
ScreenModuleEditorView "ControlMotor-NoAUTO" 640x480
   Button "Botón_1" at 10,10 size 109x37
   Button "Botón_2" at 10,50 size 109x37
   Button "Botón_3" at 130,10 size 101x37
   Button "Botón_4" at 130,50 size 101x37
*)

(* ===== HMI "HMI_RT_1" =====

text list "Enclavamientos": 0 ''; 1 ''; 2 ''; 3 ''; 4 ''; 5 ''

ScreenModuleEditorView "Faceplate_7" 640x480
   Button "Botón_3" at 25,15 size 189x37
   Button "Botón_1" at 11,10 size 93x40
   Button "Botón_2" at 11,54 size 93x40
   IOField "Campo ES_1" at 143,19 size 84x26
   IOField "Campo ES_2" at 143,62 size 84x26
   TextField "Campo de texto_2" at 109,19 size 27x23
   TextField "Campo de texto_3" at 109,62 size 32x23
   IOField "Campo ES_3" at 143,19 size 84x26
   IOField "Campo ES_4" at 143,62 size 84x26
   TextField "Campo de texto_4" at 109,19 size 27x23
   TextField "Campo de texto_5" at 109,62 size 32x23
   TextField "Campo de texto_1" at 10,31 size 97x40
*)

(* ===== HMI "HMI_RT_1" =====

text list "Enclavamientos": 0 ''; 1 ''; 2 ''; 3 ''; 4 ''; 5 ''

ScreenModuleEditorView "Faceplate_2" 640x480
   TextField "Campo de texto_14" at 112,50 size 40x22
   TextField "Campo de texto_13" at 112,14 size 40x22
   TextField "Campo de texto_1" at 67,18 size 125x50
   Button "Botón_1" at 11,10 size 93x32
   Button "Botón_2" at 11,46 size 93x32
   Button "Botón_3" at 136,10 size 117x32
   Button "Botón_4" at 136,46 size 117x32
   SymbolicIOField "Campo ES simbólico_2" at 158,12 size 96x27
   SymbolicIOField "Campo ES simbólico_3" at 158,47 size 96x27
*)

(* ===== HMI "HMI_RT_1" =====

text list "EstadoMotor": 0 ''; 1 ''; 2 ''; 3 ''; 4 ''; 5 ''; 6 ''; 7 ''

ScreenModuleEditorView "ControlMotor-NoAUTO" 640x480
   Button "Botón_1" at 10,10 size 109x37
   Button "Botón_2" at 10,50 size 109x37
   Button "Botón_3" at 130,10 size 101x37
   Button "Botón_4" at 130,50 size 101x37
*)

(* ===== HMI "HMI_RT_1" =====

ScreenModuleEditorView "Faceplate_4" 640x480
   TextField "Campo de texto_14" at 117,50 size 25x22
   TextField "Campo de texto_13" at 119,14 size 23x22
   IOField "Campo ES_9" at 147,48 size 83x29
   IOField "Campo ES_8" at 147,12 size 83x29
   Button "Botón_1" at 10,10 size 93x32
   Button "Botón_2" at 10,46 size 93x32
   Button "Botón_3" at 122,10 size 109x32
   Button "Botón_4" at 122,46 size 109x32
*)

(* ===== HMI "HMI_RT_1" =====

ScreenModuleEditorView "Faceplate_1" 640x480
   TextField "Campo de texto_14" at 117,50 size 25x22
   TextField "Campo de texto_13" at 119,14 size 23x22
   IOField "Campo ES_9" at 147,48 size 83x29
   IOField "Campo ES_8" at 147,12 size 83x29
   Button "Botón_1" at 10,10 size 93x32
   Button "Botón_2" at 10,46 size 93x32
   Button "Botón_3" at 122,10 size 109x32
   Button "Botón_4" at 122,46 size 109x32
*)

(* ===== HMI "HMI_RT_1" =====

ScreenModuleEditorView "Faceplate_1" 640x480
   TextField "Campo de texto_14" at 118,50 size 25x22
   TextField "Campo de texto_13" at 120,14 size 23x22
   TextField "Campo de texto_1" at 59,18 size 125x50
   IOField "Campo ES_9" at 148,48 size 83x29
   IOField "Campo ES_8" at 148,12 size 83x29
   Button "Botón_1" at 11,10 size 93x32
   Button "Botón_2" at 11,46 size 93x32
   Button "Botón_3" at 123,10 size 109x32
   Button "Botón_4" at 123,46 size 109x32
*)

(* ===== HMI "HMI_RT_1" =====

text list "Enclavamientos": 0 ''; 1 ''; 2 ''; 3 ''; 4 ''; 5 ''

ScreenModuleEditorView "Faceplate_10" 640x480
   Button "Botón_3" at 38,10 size 189x37
   Button "Botón_1" at 38,10 size 93x40
   Button "Botón_2" at 133,10 size 93x40
   IOField "Campo ES_1" at 44,75 size 84x26
   IOField "Campo ES_2" at 44,110 size 84x26
   TextField "Campo de texto_2" at 10,75 size 27x23
   TextField "Campo de texto_3" at 10,110 size 32x23
   IOField "Campo ES_3" at 140,75 size 84x26
   IOField "Campo ES_4" at 140,110 size 84x26
   TextField "Campo de texto_4" at 60,51 size 45x23
   TextField "Campo de texto_5" at 146,51 size 71x23
   IOField "Campo ES_5" at 44,75 size 84x26
   IOField "Campo ES_6" at 44,110 size 84x26
   IOField "Campo ES_7" at 140,75 size 84x26
   IOField "Campo ES_8" at 140,110 size 84x26
   TextField "Campo de texto_6" at 10,75 size 27x23
   TextField "Campo de texto_7" at 10,110 size 32x23
   TextField "Campo de texto_8" at 60,51 size 45x23
   TextField "Campo de texto_9" at 146,51 size 71x23
   TextField "Campo de texto_1" at 77,12 size 108x42
*)

(* ===== HMI "HMI_RT_1" =====

ScreenModuleEditorView "Faceplate_6" 640x480
   GraphicIOField "PlotLight_Round_GN" at 52,10 size 35x34
   GraphicIOField "PlotLight_Round_RN" at 10,10 size 34x34
   GraphicView "Visor de gráficos_1" at 52,10 size 34x34
   GraphicView "Visor de gráficos_2" at 53,10 size 34x34
*)

(* ===== HMI "HMI_RT_1" =====

ScreenModuleEditorView "Faceplate_1" 640x480
   Button "Botón_1" at 10,10 size 93x32
   Button "Botón_2" at 10,46 size 93x32
   Button "Botón_3" at 122,10 size 109x32
   Button "Botón_4" at 122,46 size 109x32
*)

(* ===== HMI "HMI_RT_1" =====
connection "Conexión-PLC_2": ETHERNET, SIMATIC S7 300/400 MPI
connection "Conexión-SentronPac_": ETHERNET, MODBUS_TCP

HMI tags "Tabla de variables estándar"
   "IndR6" : Bool, 100 ms
   "IndVparp6" : Bool, 1 s
   "Auto6" : Bool, 1 s
   "PanMCH6" : Bool, 1 s
   "LimSUP6" : Real, 1 s
   "LimINF6" : Real, 1 s
   "VCMP6" : Int, 1 s
   "IncP6" : Bool, 100 ms
   "DecP6" : Bool, 1 s
   "SPONF6" : Real, 1 s
   "SPOFFF6" : Real, 1 s
   "ForzarMarcha6" : Bool, 1 s
   "ForzarParada6" : Bool, 1 s
   "ForzandoMarcha6" : Bool, 1 s
   "SPON6" : Real, 1 s
   "SPOFF6" : Real, 1 s
   "AnimMenuMC006" : Int, 1 s
   "MantMC006" : Bool, 1 s
   "MarchaOK6" : Bool, 1 s
   "MarchaMC006" : Bool, 1 s
   "ParadaMC006" : Bool, 1 s
   "HORAS6" : DInt, 1 s
   "MIN6" : Int, 1 s
   "AnimMotorMC006" : Byte, 1 s
   "EV6" : Bool, 1 s
   "EnclavCompAltaConFlujostato" : Bool = PLC "EnclavCompAltaConFlujostato", 1 s
   "ProxMantMC001_1" : DInt = PLC "ProxMantMC001_1", 1 s
   "ProxMantMC001_2" : DInt = PLC "ProxMantMC001_2", 1 s
   "Varios_UltimoMantMC001_1" : DInt, 1 s
   "Varios_UltimoMantMC001_2" : DInt, 1 s
   "ProxMantMC002_1" : DInt = PLC "ProxMantMC002_1", 1 s
   "ProxMantMC002_2" : DInt = PLC "ProxMantMC002_2", 1 s
   "ProxMantMC003_1" : DInt = PLC "ProxMantMC003_1", 1 s
   "ProxMantMC003_2" : DInt = PLC "ProxMantMC003_2", 1 s
   "ProxMantMC004_1" : DInt = PLC "ProxMantMC004_1", 1 s
   "ProxMantMC004_2" : DInt = PLC "ProxMantMC004_2", 1 s
   "ProxMantMC005_1" : DInt = PLC "ProxMantMC005_1", 1 s
   "ProxMantMC005_2" : DInt = PLC "ProxMantMC005_2", 1 s
   "ProxMantMC006_1" : DInt = PLC "ProxMantMC006_1", 1 s
   "ProxMantMC006_2" : DInt = PLC "ProxMantMC006_2", 1 s
   "Varios_UltimoMantMC002_1" : DInt, 1 s
   "Varios_UltimoMantMC002_2" : DInt, 1 s
   "Varios_UltimoMantMC003_1" : DInt, 1 s
   "Varios_UltimoMantMC003_2" : DInt, 1 s
   "Varios_UltimoMantMC004_1" : DInt, 1 s
   "Varios_UltimoMantMC004_2" : DInt, 1 s
   "Varios_UltimoMantMC005_1" : DInt, 1 s
   "Varios_UltimoMantMC005_2" : DInt, 1 s
   "Varios_UltimoMantMC006_1" : DInt, 1 s
   "Varios_UltimoMantMC006_2" : DInt, 1 s
   "Varios_HorasMantMC001_1" : DInt, 1 s
   "Varios_HorasMantMC006_1" : DInt, 1 s
   "Varios_HorasMantMC006_2" : DInt, 1 s
   "Varios_HorasMantMC002_1" : DInt, 1 s
   "Varios_HorasMantMC001_2" : DInt, 1 s
   "Varios_HorasMantMC002_2" : DInt, 1 s
   "Varios_HorasMantMC004_1" : DInt, 1 s
   "Varios_HorasMantMC004_2" : DInt, 1 s
   "Varios_HorasMantMC005_1" : DInt, 1 s
   "Varios_HorasMantMC005_2" : DInt, 1 s
   "Varios_HorasMantMC003_1" : DInt, 1 s
   "Varios_HorasMantMC003_2" : DInt, 1 s
   "EstadoMantMC003" : Byte = PLC "EstadoMantMC003", 1 s
   "EstadoMantMC005" : Byte = PLC "EstadoMantMC005", 1 s
   "EstadoMantMC004" : Byte = PLC "EstadoMantMC004", 1 s
   "EstadoMantMC002" : Byte = PLC "EstadoMantMC002", 1 s
   "EstadoMantMC001" : Byte = PLC "EstadoMantMC001", 1 s
   "EstadoMantMC006" : Byte = PLC "EstadoMantMC006", 1 s
   "LimiteMantMC001_1" : Bool = PLC "LimiteMantMC001_1", 1 s
   "LimiteMantMC001_2" : Bool = PLC "LimiteMantMC001_2", 1 s
   "LimiteMantMC002_1" : Bool = PLC "LimiteMantMC002_1", 1 s
   "LimiteMantMC002_2" : Bool = PLC "LimiteMantMC002_2", 1 s
   "LimiteMantMC003_1" : Bool = PLC "LimiteMantMC003_1", 1 s
   "LimiteMantMC003_2" : Bool = PLC "LimiteMantMC003_2", 1 s
   "LimiteMantMC004_1" : Bool = PLC "LimiteMantMC004_1", 1 s
   "LimiteMantMC004_2" : Bool = PLC "LimiteMantMC004_2", 1 s
   "LimiteMantMC005_1" : Bool = PLC "LimiteMantMC005_1", 1 s
   "LimiteMantMC005_2" : Bool = PLC "LimiteMantMC005_2", 1 s
   "LimiteMantMC006_1" : Bool = PLC "LimiteMantMC006_1", 1 s
   "LimiteMantMC006_2" : Bool = PLC "LimiteMantMC006_2", 1 s
   "Varios_HorasMantMS050" : DInt, 1 s
   "Varios_HorasMantMS051" : DInt, 1 s
   "Varios_HorasMantMS052" : DInt, 1 s
   "Varios_HorasMantMS053" : DInt, 1 s
   "HorasSecAlta_HMMS050" : DInt, 1 s
   "HorasSecAlta_HMMS051" : DInt, 1 s
   "HorasSecAlta_HMMS052" : DInt, 1 s
   "HorasSecAlta_HMMS053" : DInt, 1 s
   "Varios_UltimoMantMS050" : DInt, 1 s
   "HorasSecAlta_MMMS050" : Int, 1 s
   "ProxMantMS050" : DInt = PLC "ProxMantMS050", 1 s
   "Varios_UltimoMantMS051" : DInt, 1 s
   "ProxMantMS051" : DInt = PLC "ProxMantMS051", 1 s
   "HorasSecAlta_MMMS051" : Int, 1 s
   "Varios_UltimoMantMS052" : DInt, 1 s
   "ProxMantMS052" : DInt = PLC "ProxMantMS052", 1 s
   "HorasSecAlta_MMMS052" : Int, 1 s
   "Varios_UltimoMantMS053" : DInt, 1 s
   "ProxMantMS053" : DInt = PLC "ProxMantMS053", 1 s
   "HorasSecAlta_MMMS053" : Int, 1 s
   "LimiteMantMS051" : Bool = PLC "LimiteMantMS051", 1 s
   "LimiteMantMS053" : Bool = PLC "LimiteMantMS053", 1 s
   "LimiteMantMS052" : Bool = PLC "LimiteMantMS052", 1 s
   "LimiteMantMS050" : Bool = PLC "LimiteMantMS050", 1 s
   "Varios_HorasMantMC060_1" : DInt, 1 s
   "Varios_HorasMantMC060_2" : DInt, 1 s
   "Varios_HorasMantMC060_3" : DInt, 1 s
   "Varios_HorasMantMC060_4" : DInt, 1 s
   "Varios_UltimoMantMC060_5" : DInt, 1 s
   "Varios_UltimoMantMC062_1" : DInt, 1 s
   "Varios_HorasMantMC061_1" : DInt, 1 s
   "Varios_HorasMantMC061_2" : DInt, 1 s
   "Varios_HorasMantMC061_3" : DInt, 1 s
   "Varios_HorasMantMC061_4" : DInt, 1 s
   "Varios_HorasMantMC061_5" : DInt, 1 s
   "Varios_HorasMantMC062_1" : DInt, 1 s
   "Varios_HorasMantMC062_2" : DInt, 1 s
   "Varios_HorasMantMC062_3" : DInt, 1 s
   "Varios_HorasMantMC062_4" : DInt, 1 s
   "Varios_HorasMantMC062_5" : DInt, 1 s
   "Varios_HorasMantMC063_1" : DInt, 1 s
   "Varios_HorasMantMC063_2" : DInt, 1 s
   "Varios_HorasMantMC063_3" : DInt, 1 s
   "Varios_HorasMantMC063_4" : DInt, 1 s
   "Varios_HorasMantMC063_5" : DInt, 1 s
   "Varios_HorasMantMC064_1" : DInt, 1 s
   "Varios_HorasMantMC064_2" : DInt, 1 s
   "Varios_HorasMantMC064_3" : DInt, 1 s
   "Varios_HorasMantMC064_4" : DInt, 1 s
   "Varios_HorasMantMC064_5" : DInt, 1 s
   "Varios_HorasMantMS054_1" : DInt, 1 s
   "Varios_HorasMantMS054_2" : DInt, 1 s
   "Varios_UltimoMantMS055_1" : DInt, 1 s
   "Varios_HorasMantMS055_2" : DInt, 1 s
   "HorasCmpBaja_HMMC060" : DInt, 1 s
   "HorasCmpBaja_MMMC060" : Int, 1 s
   "Varios_UltimoMantMC060_1" : DInt, 1 s
   "ProxMantMC060_1" : DInt = PLC "ProxMantMC060_1", 1 s
   "ProxMantMC060_2" : DInt = PLC "ProxMantMC060_2", 1 s
   "ProxMantMC060_3" : DInt = PLC "ProxMantMC060_3", 1 s
   "ProxMantMC060_4" : DInt = PLC "ProxMantMC060_4", 1 s
   "ProxMantMC060_5" : DInt = PLC "ProxMantMC060_5", 1 s
   "Varios_UltimoMantMC060_2" : DInt, 1 s
   "Varios_UltimoMantMC060_3" : DInt, 1 s
   "Varios_UltimoMantMC060_4" : DInt, 1 s
   "HorasCmpBaja_HMMC061" : DInt, 1 s
   "ProxMantMC061_1" : DInt = PLC "ProxMantMC061_1", 1 s
   "ProxMantMC061_3" : DInt = PLC "ProxMantMC061_3", 1 s
   "ProxMantMC061_4" : DInt = PLC "ProxMantMC061_4", 1 s
   "ProxMantMC061_2" : DInt = PLC "ProxMantMC061_2", 1 s
   "ProxMantMC061_5" : DInt = PLC "ProxMantMC061_5", 1 s
   "Varios_UltimoMantMC061_1" : DInt, 1 s
   "Varios_UltimoMantMC061_2" : DInt, 1 s
   "Varios_UltimoMantMC061_3" : DInt, 1 s
   "Varios_UltimoMantMC061_4" : DInt, 1 s
   "Varios_UltimoMantMC061_5" : DInt, 1 s
   "HorasCmpBaja_MMMC061" : Int, 1 s
   "HorasCmpBaja_HMMC062" : DInt, 1 s
   "HorasCmpBaja_MMMC062" : Int, 1 s
   "ProxMantMC062_1" : DInt = PLC "ProxMantMC062_1", 1 s
   "ProxMantMC062_2" : DInt = PLC "ProxMantMC062_2", 1 s
   "ProxMantMC062_3" : DInt = PLC "ProxMantMC062_3", 1 s
   "ProxMantMC062_4" : DInt = PLC "ProxMantMC062_4", 1 s
   "ProxMantMC062_5" : DInt = PLC "ProxMantMC062_5", 1 s
   "Varios_UltimoMantMC062_5" : DInt, 1 s
   "Varios_UltimoMantMC062_3" : DInt, 1 s
   "Varios_UltimoMantMC062_2" : DInt, 1 s
   "HorasCmpBaja_HMMC063" : DInt, 1 s
   "HorasCmpBaja_MMMC063" : Int, 1 s
   "ProxMantMC063_1" : DInt = PLC "ProxMantMC063_1", 1 s
   "ProxMantMC063_2" : DInt = PLC "ProxMantMC063_2", 1 s
   "ProxMantMC063_3" : DInt = PLC "ProxMantMC063_3", 1 s
   "ProxMantMC063_4" : DInt = PLC "ProxMantMC063_4", 1 s
   "ProxMantMC063_5" : DInt = PLC "ProxMantMC063_5", 1 s
   "HorasCmpBaja_HMMC064" : DInt, 1 s
   "Varios_UltimoMantMC063_1" : DInt, 1 s
   "Varios_UltimoMantMC063_2" : DInt, 1 s
   "Varios_UltimoMantMC063_3" : DInt, 1 s
   "Varios_UltimoMantMC063_4" : DInt, 1 s
   "Varios_UltimoMantMC063_5" : DInt, 1 s
   "HorasCmpBaja_MMMC064" : Int, 1 s
   "ProxMantMC064_1" : DInt = PLC "ProxMantMC064_1", 1 s
   "ProxMantMC064_2" : DInt = PLC "ProxMantMC064_2", 1 s
   "ProxMantMC064_3" : DInt = PLC "ProxMantMC064_3", 1 s
   "ProxMantMC064_4" : DInt = PLC "ProxMantMC064_4", 1 s
   "ProxMantMC064_5" : DInt = PLC "ProxMantMC064_5", 1 s
   "Varios_UltimoMantMC064_1" : DInt, 1 s
   "Varios_UltimoMantMC064_5" : DInt, 1 s
   "Varios_UltimoMantMC064_2" : DInt, 1 s
   "Varios_UltimoMantMC064_3" : DInt, 1 s
   "Varios_UltimoMantMC064_4" : DInt, 1 s
   "LimiteMantMC060_1" : Bool = PLC "LimiteMantMC060_1", 1 s
   "LimiteMantMC060_2" : Bool = PLC "LimiteMantMC060_2", 1 s
   "LimiteMantMC060_3" : Bool = PLC "LimiteMantMC060_3", 1 s
   "LimiteMantMC060_4" : Bool = PLC "LimiteMantMC060_4", 1 s
   "LimiteMantMC060_5" : Bool = PLC "LimiteMantMC060_5", 1 s
   "EstadoMantMC060" : Byte = PLC "EstadoMantMC060", 1 s
   "EstadoMantMC061" : Byte = PLC "EstadoMantMC061", 1 s
   "EstadoMantMC062" : Byte = PLC "EstadoMantMC062", 1 s
   "EstadoMantMC063" : Byte = PLC "EstadoMantMC063", 1 s
   "EstadoMantMC064" : Byte = PLC "EstadoMantMC064", 1 s
   "HorasSecBaja_HMMS054" : DInt, 1 s
   "HorasSecBaja_MMMS054" : Int, 1 s
   "ProxMantMS054_1" : DInt = PLC "ProxMantMS054_1", 1 s
   "ProxMantMS054_2" : DInt = PLC "ProxMantMS054_2", 1 s
   "Varios_UltimoMantMS054_1" : DInt, 1 s
   "Varios_UltimoMantMS054_2" : DInt, 1 s
   "EstadoMantSecBaja" : Byte = PLC "EstadoMantSecBaja", 1 s
   "LimiteMantMS054_1" : Bool = PLC "LimiteMantMS054_1", 1 s
   "LimiteMantMS054_2" : Bool = PLC "LimiteMantMS054_2", 1 s
   "LimiteMantMS055_1" : Bool = PLC "LimiteMantMS055_1", 1 s
   "LimiteMantMS055_2" : Bool = PLC "LimiteMantMS055_2", 1 s
   "HorasSecBaja_HMMS055" : DInt, 1 s
   "HorasSecBaja_MMMS055" : Int, 1 s
   "ProxMantMS055_1" : DInt = PLC "ProxMantMS055_1", 1 s
   "ProxMantMS055_2" : DInt = PLC "ProxMantMS055_2", 1 s
   "Varios_UltimoMantMS055_2" : DInt, 1 s
   "Varios_HorasMantBost1" : DInt, 1 s
   "Varios_HorasMantBost2" : DInt, 1 s
   "ProxMantBoost1" : DInt = PLC "ProxMantBoost1", 1 s
   "ProxMantBoost2" : DInt = PLC "ProxMantBoost2", 1 s
   "Varios_UltimoMantBoost1" : DInt, 1 s
   "Varios_UltimoMantBoost2" : DInt, 1 s
   "LimiteMantBoost1" : Bool = PLC "LimiteMantBoost1", 1 s
   "LimiteMantBoost2" : Bool = PLC "LimiteMantBoost2", 1 s
   "DBParamCmpALTA-MTA_TempCritEnclav" : Real, 1 s
   "EnclavCompAltaPorTemp" : Bool = PLC "EnclavCompAltaPorTemp", 1 s
   "NumeroCompresor" : Int, internal
   "EstadoRegistro" : Bool, internal

HMI tags "Tabla de variables estándar_1"
   "MC066_STD" : , 1 s
   "MV031_STD" : , 1 s
   "MV032_STD" : , 1 s
   "MV030_STD" : , 1 s
   "DIP_1" : , internal
   "MP016_STD" : , 1 s
   "MC004_STD" : , 1 s
   "MP013_STD" : , 1 s
   "MV033_STD" : , 1 s
   "MC001_STD" : , 1 s
   "MC060_STD" : , 1 s
   "MC002_STD" : , 1 s
   "MP012_STD" : , 1 s
   "MC065_STD" : , 1 s
   "MS051_STD" : , 1 s
   "MC006_STD" : , 1 s
   "MP011_STD" : , 1 s
   "Iluminati_STD" : , 1 s
   "MC064_STD" : , 1 s
   "MS052_STD" : , 1 s
   "MT010_STD" : , 1 s
   "MS053_STD" : , 1 s
   "MP019_STD" : , 1 s
   "MC005_STD" : , 1 s
   "MC061_STD" : , 1 s
   "MV034_STD" : , 1 s
   "MC063_STD" : , 1 s
   "MP015_STD" : , 1 s
   "MT007_STD" : , 1 s
   "MS055_STD" : , 1 s
   "MP018_STD" : , 1 s
   "MP014_STD" : , 1 s
   "MS054_STD" : , 1 s
   "MS050_STD" : , 1 s
   "MP010_STD" : , 1 s
   "MT008_STD" : , 1 s
   "MT009_STD" : , 1 s
   "MC003_STD" : , 1 s
   "MC062_STD" : , 1 s
   "EB5" : Word, 1 s
   "EB7" : Word, 1 s
   "EB4" : Word, 1 s
   "EW8" : Word, 1 s
   "ACK_ALARMA_2" : Int, 1 s
   "MP020_STD" : Word, 1 s
   "MP021_STD" : Word, 1 s
   "MP022_STD" : Word, 1 s
   "CERO" : Bool, 1 s
   "UNO" : Bool, 1 s
   "IndCh" : Bool, 1 s
   "IndTrCh" : Bool, 1 s
   "IndCmpBaja" : Bool, 1 s
   "IndSecBaja" : Bool, 1 s
   "IndCmpAlta" : Bool, 1 s
   "IndSecAlta" : Bool, 1 s
   "IndTrCav" : Bool, 1 s
   "AnularSirena?" : Bool, internal
   "HorasBoost1" : DInt, 1 s
   "HorasBoost2" : DInt, 1 s
   "BoostPrHoras" : Bool, 1 s
   "BoostInvP" : Bool, 1 s
   "PrioridadBoost1" : Int, 1 s
   "PrioridadBoost2" : Int, 1 s
   "BoostInvPMan" : Bool, 1 s
   "min_boost1" : Int, 1 s
   "SegsBoost1" : Int, 1 s
   "SegsBoost" : Int, 1 s
   "MinBoost2" : Int, 1 s
   "FT1_AGUA" : Bool = PLC "FT1_AGUA", 1 s

HMI tags "AlarmasMTA"
   "AlarmasWord0" : Int, 1 s
   "AlarmasWord1" : Int, 1 s
   "AlarmasWord2" : Int, 1 s
   "AlarmasWord3" : Int, 1 s
   "AlarmasWord4" : Int, 1 s
   "AlarmasWord5" : Int, 1 s
   "AlarmasWord6" : Int, 1 s
   "AlarmasWord7" : Int, 1 s
   "AlarmasWord8" : Int, 1 s
   "Rec0" : Int, 1 s
   "Rec1" : Int, 1 s
   "Rec2" : Int, 1 s
   "Rec3" : Int, 1 s
   "Rec4" : Int, 1 s
   "Rec5" : Int, 1 s
   "Rec6" : Int, 1 s
   "Rec7" : Int, 1 s
   "Rec8" : Int, 1 s
   "AlarmasWord9" : Int, 1 s
   "AlarmasWord10" : Int, 1 s
   "AlarmasWord11" : Int, 1 s
   "AlarmasWord12" : Int, 1 s
   "AlarmasWord13" : Int, 1 s
   "AlarmasWord14" : Int, 1 s
   "Rec9" : Int, 1 s
   "Rec10" : Int, 1 s
   "Rec11" : Int, 1 s
   "Rec12" : Int, 1 s
   "Rec13" : Int, 1 s
   "Rec14" : Int, 1 s
   "AlarmasWord15" : Int, 1 s
   "Rec15" : Int, 1 s
   "ReconocerTODAS" : Bool, 1 s
   "EncendidoPLC" : Bool, 1 s
   "AlarmasWord16" : Int, 1 s
   "Rec16" : Int, 1 s
   "ReconocerTODAS_1" : Bool, 1 s
   "AlarmasWord18" : Int, 1 s
   "Rec18" : Int, 1 s
   "AlarmasWord19" : Int, 1 s
   "Rec19" : Int, 1 s
   "AlarmasWord20" : Int, 1 s
   "AlarmasWord21" : Int, 1 s
   "AlarmasWord22" : Int, 1 s
   "AlarmasWord23" : Int, 1 s
   "AlarmasWord24" : Int, 1 s
   "Rec20" : Int, 1 s
   "Rec21" : Int, 1 s
   "Rec22" : Int, 1 s
   "Rec23" : Int, 1 s
   "Rec24" : Int, 1 s

HMI tags "AutoTorresCav"
   "AutoV030" : Bool, 1 s
   "AutoV031" : Bool, 1 s
   "SP-OFF-V030" : Int, 1 s
   "SP-OFF-V031" : Int, 1 s
   "SP-ON-V030" : Int, 1 s
   "SP-ON-V031" : Int, 1 s

HMI tags "AutoTorresChillers"
   "AutoV001" : Bool, 1 s
   "AutoV002" : Bool, 1 s
   "AutoV003" : Bool, 1 s
   "SP-ON-V001" : Int, 1 s
   "SP-ON-V002" : Int, 1 s
   "SP-ON-V003" : Int, 1 s
   "SP-OFF-V001" : Int, 1 s
   "SP-OFF-V002" : Int, 1 s
   "SP-OFF-V003" : Int, 1 s
   "TemperaturatorresCH" : Real, 1 s

HMI tags "Booster"
   "AlarmaBooster" : Bool, 1 s
   "Booster_ModoManten" : Bool, 1 s
   "Booster_ModoManual" : Bool, 1 s
   "Booster_ModoAutoma" : Bool, 1 s
   "Booster_PlsManten" : Bool, 1 s
   "Booster_PlsManual" : Bool, 1 s
   "Booster_PlsAutoma" : Bool, 1 s
   "AnimaMotBooster" : Byte, 1 s
   "BoosterOrdMarcha" : Bool, 1 s
   "Booster_Conf_Marcha" : Bool, 1 s
   "Booster_Presost_Ctrl" : Bool, 1 s
   "Booster_Presost_PA" : Bool, 1 s
   "Booster_Habilitacion" : Bool, 1 s
   "Booster2_Conf_Marcha" : Bool, 1 s
   "Booster2_Habilitacion" : Bool, 1 s
   "Booster2_ModoAutoma" : Bool, 1 s
   "Booster2_ModoManten" : Bool, 1 s
   "Booster2_ModoManual" : Bool, 1 s
   "Booster2_PlsAutoma" : Bool, 1 s
   "Booster2_PlsManten" : Bool, 1 s
   "Booster2_PlsManual" : Bool, 1 s
   "AnimaMotBooster2" : Byte, 1 s
   "Booster2OrdMarcha" : Bool, 1 s
   "TiempoAyudaON" : Int, 1 s
   "TiempoAyudaOFF" : Int, 1 s
   "DifHorINVBoost" : DInt, 1 s
   "LimArrBoostPrio2" : Real, 1 s
   "LimArrBoostPrio1" : Real, 1 s
   "LimParBoostPrio2" : Real, 1 s
   "LimParBoostPrio1" : Real, 1 s
   "Presión_Actual_Boosters" : Real, 1 s
   "Ctrl_Analógico" : Bool, 1 s
   "Ver_Config" : Bool, internal
   "CotaSupPresAna" : Real, 1 s

HMI tags "CFG-Analog-MTA"
   "PresiónALTA" : Real, 1 s
   "PresiónBAJA" : Real, 1 s
   "TempCAV" : Real, 1 s
   "TempCH" : Real, 1 s
   "CFG-ALtaHH" : Real, 1 s
   "CFG-ALtaH" : Real, 1 s
   "CFG-ALtaL" : Real, 1 s
   "CFG-ALtaLL" : Real, 1 s
   "CFG-BajaHH" : Real, 1 s
   "CFG-BajaH" : Real, 1 s
   "CFG-BajaL" : Real, 1 s
   "CFG-BajaLL" : Real, 1 s
   "LO_potencia" : Real, 1 s
   "HI_caudal" : Real, 1 s
   "LO_caudal" : Real, 1 s
   "HI_potencia" : Real, 1 s
   "Caudal" : Real, 1 s
   "Potencia" : Real, 1 s

HMI tags "ChillersMTA"
   "HabMT007" : Bool, 1 s
   "HabMT008" : Bool, 1 s
   "HabMT009" : Bool, 1 s
   "HabMT010" : Bool, 1 s
   "DesMT007" : Bool, 1 s
   "DesMT008" : Bool, 1 s
   "DesMT009" : Bool, 1 s
   "DesMT010" : Bool, 1 s
   "MarchaMT007" : Bool, 1 s
   "MarchaMT008" : Bool, 1 s
   "MarchaMT009" : Bool, 1 s
   "MarchaMT010" : Bool, 1 s
   "ParadaMT007" : Bool, 1 s
   "ParadaMT008" : Bool, 1 s
   "ParadaMT009" : Bool, 1 s
   "ParadaMT010" : Bool, 1 s
   "Habilitación-CH-SOP-GR" : Bool, 1 s
   "Habilitación-CH-SOP-CH" : Bool, 1 s
   "Habilitación-CH-ENV-GR" : Bool, 1 s
   "Habilitación-CH-ENV-CH" : Bool, 1 s
   "Alarma1-CH-SOP-GR" : Bool, 1 s
   "Alarma2-CH-SOP-GR" : Bool, 1 s
   "RUN-CH-SOP-GR" : Bool, 1 s
   "MAX-CH-SOP-GR" : Bool, 1 s
   "AnimaciónMT007" : Byte, 1 s
   "AnimaciónMT008" : Byte, 1 s
   "AnimaciónMT009" : Byte, 1 s
   "AnimaciónMT010" : Byte, 1 s
   "AnimaciónMP010" : Byte, 1 s
   "AnimaciónMP011" : Byte, 1 s
   "AnimaciónMP012" : Byte, 1 s
   "AnimaciónMP013" : Byte, 1 s
   "HabMP010" : Bool, 1 s
   "HabMP011" : Bool, 1 s
   "HabMP012" : Bool, 1 s
   "HabMP013" : Bool, 1 s
   "HabMP018" : Bool, 1 s
   "HabMP019" : Bool, 1 s
   "DesMP010" : Bool, 1 s
   "DesMP011" : Bool, 1 s
   "DesMP012" : Bool, 1 s
   "DesMP013" : Bool, 1 s
   "DesMP018" : Bool, 1 s
   "DesMP019" : Bool, 1 s
   "MarchaMP010" : Bool, 1 s
   "MarchaMP011" : Bool, 1 s
   "MarchaMP012" : Bool, 1 s
   "MarchaMP013" : Bool, 1 s
   "MarchaMP018" : Bool, 1 s
   "MarchaMP019" : Bool, 1 s
   "ParadaMP010" : Bool, 1 s
   "ParadaMP011" : Bool, 1 s
   "ParadaMP012" : Bool, 1 s
   "ParadaMP013" : Bool, 1 s
   "ParadaMP018" : Bool, 1 s
   "ParadaMP019" : Bool, 1 s
   "AnimaciónMP018" : Byte, 1 s
   "AnimaciónMP019" : Byte, 1 s
   "DesV001" : Bool, 1 s
   "DesV002" : Bool, 1 s
   "HabV001" : Bool, 1 s
   "HabV002" : Bool, 1 s
   "MarchaV001" : Bool, 1 s
   "MarchaV002" : Bool, 1 s
   "ParadaV001" : Bool, 1 s
   "ParadaV002" : Bool, 1 s
   "AnimaciónV001" : Byte, 1 s
   "AnimaciónV002" : Byte, 1 s
   "VentiladoresMTA" : Bool, internal
   "MAX-CH-ENV-GR" : Bool, 1 s
   "RUN-CH-ENV-GR" : Bool, 1 s
   "Alarma2-CH-ENV-GR" : Bool, 1 s
   "Alarma1-CH-ENV-GR" : Bool, 1 s
   "SirenaM1" : Bool, 1 s
   "SirenaM2" : Bool, 1 s
   "SirenaM3" : Bool, 1 s
   "SirenaM4" : Bool, 1 s
   "AnimaciónV003" : Byte, 1 s
   "HabV003" : Bool, 1 s
   "DesV003" : Bool, 1 s
   "MarchaV003" : Bool, 1 s
   "ParadaV003" : Bool, 1 s
   "BombaTorreON" : Bool, 1 s
   "SirenaM5" : Bool, 1 s
   "SirenaChillers" : Bool, 1 s
   "SirenaM6" : Bool, 1 s
   "SirenaM7" : Bool, 1 s
   "SirenaM8" : Bool, 1 s
   "SirenaM9" : Bool, 1 s
   "SirenaM10" : Bool, 1 s
   "AlarmaNueva" : Bool, 1 s
   "AlarmaPresente" : Bool, 1 s
   "SinAlarmas" : Bool, 1 s
   "AlarmaAceite-CH-ENV-CH" : Bool, 1 s
   "AlarmaTemp-CH-ENV-CH" : Bool, 1 s
   "RUN-CH-ENV-CH" : Bool, 1 s
   "VerCh1MTA" : Bool, internal
   "VerCh2MTA" : Bool, internal
   "VerCh3MTA" : Bool, internal
   "VerCh4MTA" : Bool, internal
   "AlarmaPRUEBA" : DWord, 1 s
   "Presosato" : Bool, 1 s
   "CH-SOP-CH-CTC1ON" : Bool, 1 s
   "CH-SOP-CH-CTC2ON" : Bool, 1 s
   "CH-SOP-CH-TERM1" : Bool, 1 s
   "CH-SOP-CH-TERM2" : Bool, 1 s
   "CH-ENV-CH-ACT" : Bool, 1 s
   "CH-ENV-CH-TEMP" : Bool, 1 s
   "CH-ENV-CH-TERM" : Bool, 1 s
   "CH-ENV-CH-RUN" : Bool, 1 s
   "BombaTorreON2" : Bool, 1 s
   "HabV001(1)" : Bool, 1 s
   "HabV002(1)" : Bool, 1 s
   "HabV003(1)" : Bool, 1 s
   "HabV4" : Bool, 1 s
   "MarchaV001(1)" : Bool, 1 s
   "MarchaV002(1)" : Bool, 1 s
   "MarchaV003(1)" : Bool, 1 s
   "ParadaV001(1)" : Bool, 1 s
   "ParadaV002(1)" : Bool, 1 s
   "ParadaV003(1)" : Bool, 1 s
   "AnimaMenuV001" : Int, 1 s
   "AnimaMenuV002" : Int, 1 s
   "AnimaMenuV003" : Int, 1 s
   "DeshV001" : Bool, 1 s
   "DeshV002" : Bool, 1 s
   "DeshV003" : Bool, 1 s

HMI tags "CompBajaMTA"
   "HabilitaciónMC060" : Bool, 1 s
   "HabilitaciónMC061" : Bool, 1 s
   "HabilitaciónMC062" : Bool, 1 s
   "HabilitaciónMC063" : Bool, 1 s
   "HabilitaciónMC064" : Bool, 1 s
   "HabilitaciónMC065" : Bool, 1 s
   "DeshabilitaciónMC060" : Bool, 1 s
   "DeshabilitaciónMC061" : Bool, 1 s
   "DeshabilitaciónMC062" : Bool, 1 s
   "DeshabilitaciónMC063" : Bool, 1 s
   "DeshabilitaciónMC064" : Bool, 1 s
   "DeshabilitaciónMC065" : Bool, 1 s
   "MarchaMC060" : Bool, 1 s
   "MarchaMC061" : Bool, 1 s
   "MarchaMC062" : Bool, 1 s
   "MarchaMC063" : Bool, 1 s
   "MarchaMC064" : Bool, 1 s
   "MarchaMC065" : Bool, 1 s
   "ParadaMC060" : Bool, 1 s
   "ParadaMC061" : Bool, 1 s
   "ParadaMC062" : Bool, 1 s
   "ParadaMC063" : Bool, 1 s
   "ParadaMC064" : Bool, 1 s
   "ParadaMC065" : Bool, 1 s
   "AnimaMC060" : Byte, 1 s
   "AnimaMC061" : Byte, 1 s
   "AnimaMC062" : Byte, 1 s
   "AnimaMC063" : Byte, 1 s
   "AnimaMC064" : Byte, 1 s
   "AnimaMC065" : Byte, 1 s
   "VerMC060" : Bool, internal
   "VerMC061" : Bool, internal
   "VerMC062" : Bool, internal
   "VerMC063" : Bool, internal
   "VerMC064" : Bool, internal
   "MantM060" : Bool, 1 s
   "MantM061" : Bool, 1 s
   "MantM062" : Bool, 1 s
   "MantM063" : Bool, 1 s
   "MantM064" : Bool, 1 s
   "AutoMC060" : Bool, 1 s
   "AutoMC061" : Bool, 1 s
   "AutoMC062" : Bool, 1 s
   "AutoMC063" : Bool, 1 s
   "AutoMC064" : Bool, 1 s
   "SponMC060" : Real, 1 s
   "SponMC061" : Real, 1 s
   "SponMC062" : Real, 1 s
   "SponMC063" : Real, 1 s
   "SponMC064" : Real, 1 s
   "SpoffMC060" : Real, 1 s
   "SpoffMC061" : Real, 1 s
   "SpoffMC062" : Real, 1 s
   "SpoffMC063" : Real, 1 s
   "SpoffMC064" : Real, 1 s
   "AnimMenuMC060" : Int, 1 s
   "AnimMenuMC061" : Int, 1 s
   "AnimMenuMC062" : Int, 1 s
   "AnimMenuMC063" : Int, 1 s
   "AnimMenuMC064" : Int, 1 s
   "HabilitarMC060" : Bool, 1 s
   "AnularSirenaCav" : Bool, 1 s
   "VerMC65" : Bool, internal

HMI tags "CompresoresAltaMTA"
   "Sop1" : Bool, 1 s
   "Sop2" : Bool, 1 s
   "Sop3" : Bool, 1 s
   "ReqSop1" : Int, 1 s
   "ReqSop2" : Int, 1 s
   "ReqSop3" : Int, 1 s
   "NinSop" : Bool, 1 s
   "VCMP1" : Int, 1 s
   "VCMP2" : Int, 1 s
   "VCMP3" : Int, 1 s
   "VCMP4" : Int, 1 s
   "VCMP5" : Int, 1 s
   "IncP1" : Bool, 100 ms
   "IncP2" : Bool, 100 ms
   "IncP3" : Bool, 100 ms
   "IncP4" : Bool, 100 ms
   "IncP5" : Bool, 100 ms
   "DecP1" : Bool, 1 s
   "DecP2" : Bool, 1 s
   "DecP3" : Bool, 1 s
   "DecP4" : Bool, 1 s
   "DecP5" : Bool, 1 s
   "PriRealCMP1" : Int, 1 s
   "PriRealCMP2" : Int, 1 s
   "PriRealCMP3" : Int, 1 s
   "PriRealCMP4" : Int, 1 s
   "PriRealCMP5" : Int, 1 s
   "Auto1" : Bool, 1 s
   "Auto2" : Bool, 1 s
   "Auto3" : Bool, 1 s
   "Auto4" : Bool, 1 s
   "Auto5" : Bool, 1 s
   "IndV1" : Bool, 100 ms
   "IndV2" : Bool, 100 ms
   "IndV3" : Bool, 100 ms
   "IndV4" : Bool, 100 ms
   "IndV5" : Bool, 100 ms
   "IndR1" : Bool, 100 ms
   "IndR2" : Bool, 100 ms
   "IndR3" : Bool, 100 ms
   "IndR4" : Bool, 100 ms
   "IndR5" : Bool, 100 ms
   "Est1" : Word, 1 s
   "Est2" : Word, 1 s
   "Est3" : Word, 1 s
   "Est4" : Word, 1 s
   "Est5" : Word, 1 s
   "LimSUP1" : Real, 1 s
   "LimSUP2" : Real, 1 s
   "LimSUP3" : Real, 1 s
   "LimSUP4" : Real, 1 s
   "LimSUP5" : Real, 1 s
   "LimINF1" : Real, 1 s
   "LimINF2" : Real, 1 s
   "LimINF3" : Real, 1 s
   "LimINF4" : Real, 1 s
   "LimINF5" : Real, 1 s
   "PresMaX" : Real, 1 s
   "Delta" : Real, 1 s
   "Hist" : Real, 1 s
   "CompReq" : Int, 1 s
   "CompReqINI" : Int, 1 s
   "AnimMenuMC001" : Int, 1 s
   "AnimMenuMC002" : Int, 1 s
   "AnimMenuMC003" : Int, 1 s
   "AnimMenuMC004" : Int, 1 s
   "AnimMenuMC005" : Int, 1 s
   "SPON1" : Real, 1 s
   "SPON2" : Real, 1 s
   "SPON3" : Real, 1 s
   "SPON4" : Real, 1 s
   "SPON5" : Real, 1 s
   "SPOFF1" : Real, 1 s
   "SPOFF2" : Real, 1 s
   "SPOFF3" : Real, 1 s
   "SPOFF4" : Real, 1 s
   "SPOFF5" : Real, 1 s
   "MantMC001" : Bool, 1 s
   "MantMC002" : Bool, 1 s
   "MantMC003" : Bool, 1 s
   "MantMC004" : Bool, 1 s
   "MantMC005" : Bool, 1 s
   "IndVparp1" : Bool, 1 s
   "IndVparp2" : Bool, 1 s
   "IndVparp3" : Bool, 1 s
   "IndVparp4" : Bool, 1 s
   "IndVparp5" : Bool, 1 s
   "TiempoenVacío" : Int, 1 s
   "TiemposinReq" : Int, 1 s
   "TiempoSop" : Int, 1 s
   "HistCRT" : Real, 1 s
   "LimINFCRT" : Real, 1 s
   "LimSUPCRT" : Real, 1 s
   "PanMCH1" : Bool, 1 s
   "PanMCH2" : Bool, 1 s
   "PanMCH3" : Bool, 1 s
   "PanMCH4" : Bool, 1 s
   "PanMCH5" : Bool, 1 s
   "MarchaMC001" : Bool, 1 s
   "MarchaMC002" : Bool, 1 s
   "MarchaMC003" : Bool, 1 s
   "MarchaMC004" : Bool, 1 s
   "MarchaMC005" : Bool, 1 s
   "ParadaMC001" : Bool, 1 s
   "ParadaMC002" : Bool, 1 s
   "ParadaMC003" : Bool, 1 s
   "ParadaMC004" : Bool, 1 s
   "ParadaMC005" : Bool, 1 s
   "AnimMotorMC001" : Byte, 1 s
   "AnimMotorMC002" : Byte, 1 s
   "AnimMotorMC003" : Byte, 1 s
   "AnimMotorMC004" : Byte, 1 s
   "AnimMotorMC005" : Byte, 1 s
   "EV1" : Bool, 1 s
   "EV2" : Bool, 1 s
   "EV3" : Bool, 1 s
   "EV4" : Bool, 1 s
   "EV5" : Bool, 1 s
   "HORAS1" : DInt, 1 s
   "HORAS2" : DInt, 1 s
   "HORAS3" : DInt, 1 s
   "HORAS4" : DInt, 1 s
   "HORAS5" : DInt, 1 s
   "MIN1" : Int, 1 s
   "MIN2" : Int, 1 s
   "MIN3" : Int, 1 s
   "MIN4" : Int, 1 s
   "MIN5" : Int, 1 s
   "MarchaOK1" : Bool, 1 s
   "MarchaOK2" : Bool, 1 s
   "MarchaOK3" : Bool, 1 s
   "MarchaOK4" : Bool, 1 s
   "MarchaOK5" : Bool, 1 s
   "ForzarMarcha1" : Bool, 1 s
   "ForzarMarcha2" : Bool, 1 s
   "ForzarMarcha3" : Bool, 1 s
   "ForzarMarcha4" : Bool, 1 s
   "ForzarMarcha5" : Bool, 1 s
   "ForzarParada1" : Bool, 1 s
   "ForzarParada2" : Bool, 1 s
   "ForzarParada3" : Bool, 1 s
   "ForzarParada4" : Bool, 1 s
   "ForzarParada5" : Bool, 1 s
   "SPONF1" : Real, 1 s
   "SPONF2" : Real, 1 s
   "SPONF3" : Real, 1 s
   "SPONF4" : Real, 1 s
   "SPONF5" : Real, 1 s
   "SPOFFF1" : Real, 1 s
   "SPOFFF2" : Real, 1 s
   "SPOFFF3" : Real, 1 s
   "SPOFFF4" : Real, 1 s
   "SPOFFF5" : Real, 1 s
   "ForzandoMarcha1" : Bool, 1 s
   "ForzandoMarcha2" : Bool, 1 s
   "ForzandoMarcha3" : Bool, 1 s
   "ForzandoMarcha4" : Bool, 1 s
   "ForzandoMarcha5" : Bool, 1 s
   "MediaCargaBellis" : Bool, 1 s
   "SPONF3b" : Real, 1 s
   "SPOFFF3b" : Real, 1 s
   "EV3b" : Bool, 1 s
   "TiempoMaxBellismedia" : Int, 1 s
   "Est6" : Int, 1 s
   "PriRealCMP6" : Int, 1 s
   "IndV6" : Bool, 1 s

HMI tags "IluminaciónMTA"
   "TiempoIluminación" : Word, 1 s
   "EncendidoPanel" : Bool, 1 s
   "ApagadoPanel" : Bool, 1 s
   "ON" : Bool, 1 s
   "MantenerON" : Bool, 1 s
   "AlarmaBoosters" : Bool, 1 s

HMI tags "SecadoresAltaMTA"
   "AnimaMS050" : Byte, 1 s
   "AnimaMS051" : Byte, 1 s
   "AnimaMS052" : Byte, 1 s
   "AnimaMS053" : Byte, 1 s
   "DeshabilitaciónMS050" : Bool, 1 s
   "DeshabilitaciónMS051" : Bool, 1 s
   "DeshabilitaciónMS052" : Bool, 1 s
   "DeshabilitaciónMS053" : Bool, 1 s
   "HabilitaciónMS050" : Bool, 1 s
   "HabilitaciónMS051" : Bool, 1 s
   "HabilitaciónMS052" : Bool, 1 s
   "HabilitaciónMS053" : Bool, 1 s
   "MantMS050" : Bool, 1 s
   "MantMS051" : Bool, 1 s
   "MantMS052" : Bool, 1 s
   "MantMS053" : Bool, 1 s
   "MarchaMS050" : Bool, 1 s
   "MarchaMS051" : Bool, 1 s
   "MarchaMS052" : Bool, 1 s
   "MarchaMS053" : Bool, 1 s
   "ParadaMS050" : Bool, 1 s
   "ParadaMS051" : Bool, 1 s
   "ParadaMS052" : Bool, 1 s
   "ParadaMS053" : Bool, 1 s
   "AnimaMenuMS050" : Int, 1 s
   "AnimaMenuMS051" : Int, 1 s
   "AnimaMenuMS052" : Int, 1 s
   "AnimaMenuMS053" : Int, 1 s
   "Enc1MS050" : Int, 1 s
   "Enc2MS050" : Int, 1 s
   "Enc1MS051" : Int, 1 s
   "Enc2MS051" : Int, 1 s
   "Enc1MS052" : Int, 1 s
   "Enc2MS052" : Int, 1 s
   "Enc1MS053" : Int, 1 s
   "Enc2MS053" : Int, 1 s
   "AutoMS050" : Bool, 1 s
   "AutoMS051" : Bool, 1 s
   "AutoMS052" : Bool, 1 s
   "AutoMS053" : Bool, 1 s

HMI tags "SecadoresBaja"
   "AnimaMS054" : Byte, 1 s
   "AnimaMS055" : Byte, 1 s
   "DeshabilitaciónMS054" : Bool, 1 s
   "DeshabilitaciónMS055" : Bool, 1 s
   "HabilitaciónMS054" : Bool, 1 s
   "HabilitaciónMS055" : Bool, 1 s
   "MarchaMS054" : Bool, 1 s
   "MarchaMS055" : Bool, 1 s
   "ParadaMS054" : Bool, 1 s
   "ParadaMS055" : Bool, 1 s
   "MantMS054" : Bool, 1 s
   "MantMS055" : Bool, 1 s
